REGION Network 3
   RUNG wire#powerrail
      Contact( "FB11_DATA_ALARM_FB_DB".PIW258.QH_ALM )
      wire#w1
      P_Trig( "DB9_P".P2 )
      S_Coil( "Tag_32" )
   END_RUNG
   RUNG wire#powerrail
      Contact( "FB11_DATA_ALARM_FB_DB".PIW258.QL_ALM )
   END_RUNG wire#w1
   // the same network as SCL:
   #_w1 := "FB11_DATA_ALARM_FB_DB".PIW258.QH_ALM OR "FB11_DATA_ALARM_FB_DB".PIW258.QL_ALM;
   #_w2 := #_w1 AND NOT "DB9_P".P2;   // rising edge
   "DB9_P".P2 := #_w1;
   IF #_w2 THEN "Tag_32" := TRUE; END_IF;
END_REGION

REGION Network 4
   RUNG wire#powerrail
      Contact( "FB11_DATA_ALARM_FB_DB".PIW260.QH_ALM )
      wire#w1
      P_Trig( "DB9_P".P3 )
      S_Coil( "Tag_32" )
   END_RUNG
   RUNG wire#powerrail
      Contact( "FB11_DATA_ALARM_FB_DB".PIW260.QL_ALM )
   END_RUNG wire#w1
   // the same network as SCL:
   #_w1 := "FB11_DATA_ALARM_FB_DB".PIW260.QH_ALM OR "FB11_DATA_ALARM_FB_DB".PIW260.QL_ALM;
   #_w2 := #_w1 AND NOT "DB9_P".P3;   // rising edge
   "DB9_P".P3 := #_w1;
   IF #_w2 THEN "Tag_32" := TRUE; END_IF;
END_REGION

REGION Network 5
   RUNG wire#powerrail
      Contact( "FB11_DATA_ALARM_FB_DB".PIW262.QH_ALM )
      wire#w1
      P_Trig( "DB9_P".P4 )
      S_Coil( "Tag_32" )
   END_RUNG
   RUNG wire#powerrail
      Contact( "FB11_DATA_ALARM_FB_DB".PIW262.QL_ALM )
   END_RUNG wire#w1
   // the same network as SCL:
   #_w1 := "FB11_DATA_ALARM_FB_DB".PIW262.QH_ALM OR "FB11_DATA_ALARM_FB_DB".PIW262.QL_ALM;
   #_w2 := #_w1 AND NOT "DB9_P".P4;   // rising edge
   "DB9_P".P4 := #_w1;
   IF #_w2 THEN "Tag_32" := TRUE; END_IF;
END_REGION

REGION Network 6
   RUNG wire#powerrail
      Contact( "FB11_DATA_ALARM_FB_DB".PIW264.QH_ALM )
      wire#w1
      P_Trig( "DB9_P".P5 )
      S_Coil( "Tag_32" )
   END_RUNG
   RUNG wire#powerrail
      Contact( "FB11_DATA_ALARM_FB_DB".PIW264.QL_ALM )
   END_RUNG wire#w1
   // the same network as SCL:
   #_w1 := "FB11_DATA_ALARM_FB_DB".PIW264.QH_ALM OR "FB11_DATA_ALARM_FB_DB".PIW264.QL_ALM;
   #_w2 := #_w1 AND NOT "DB9_P".P5;   // rising edge
   "DB9_P".P5 := #_w1;
   IF #_w2 THEN "Tag_32" := TRUE; END_IF;
END_REGION

REGION Network 7
   RUNG wire#powerrail
      Contact( "FB11_DATA_ALARM_FB_DB".PIW266.QH_ALM )
      wire#w1
      P_Trig( "DB9_P".P6 )
      S_Coil( "Tag_32" )
   END_RUNG
   RUNG wire#powerrail
      Contact( "FB11_DATA_ALARM_FB_DB".PIW266.QL_ALM )
   END_RUNG wire#w1
   // the same network as SCL:
   #_w1 := "FB11_DATA_ALARM_FB_DB".PIW266.QH_ALM OR "FB11_DATA_ALARM_FB_DB".PIW266.QL_ALM;
   #_w2 := #_w1 AND NOT "DB9_P".P6;   // rising edge
   "DB9_P".P6 := #_w1;
   IF #_w2 THEN "Tag_32" := TRUE; END_IF;
END_REGION

REGION Network 8
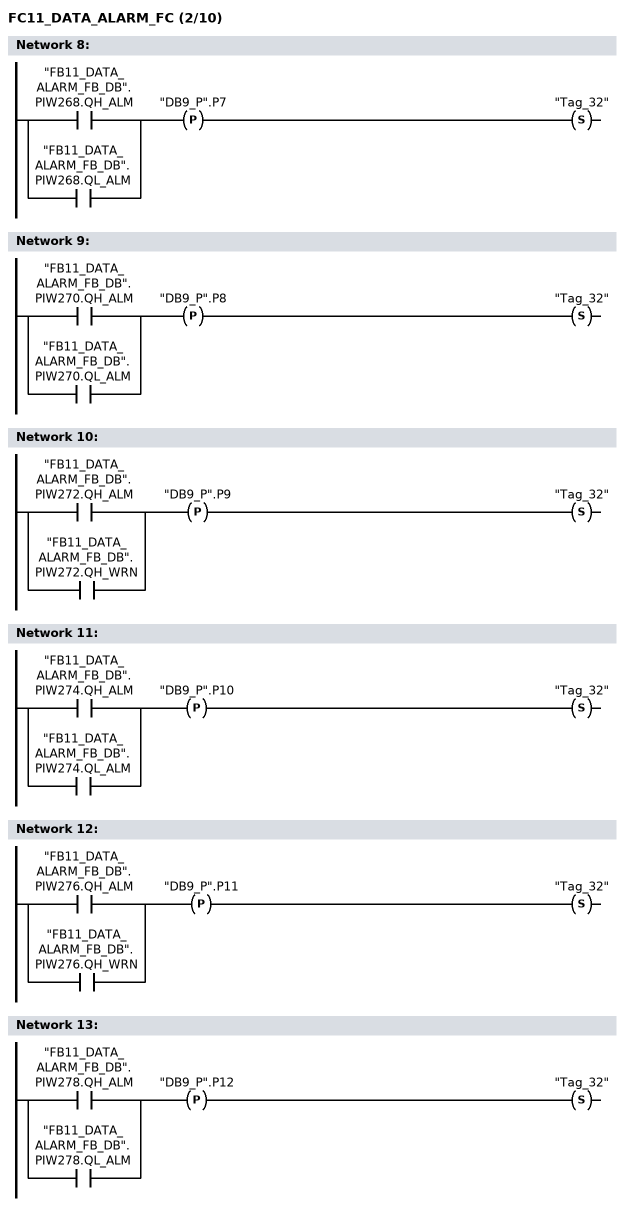
   RUNG wire#powerrail
      Contact( "FB11_DATA_ALARM_FB_DB".PIW268.QH_ALM )
      wire#w1
      P_Trig( "DB9_P".P7 )
      S_Coil( "Tag_32" )
   END_RUNG
   RUNG wire#powerrail
      Contact( "FB11_DATA_ALARM_FB_DB".PIW268.QL_ALM )
   END_RUNG wire#w1
   // the same network as SCL:
   #_w1 := "FB11_DATA_ALARM_FB_DB".PIW268.QH_ALM OR "FB11_DATA_ALARM_FB_DB".PIW268.QL_ALM;
   #_w2 := #_w1 AND NOT "DB9_P".P7;   // rising edge
   "DB9_P".P7 := #_w1;
   IF #_w2 THEN "Tag_32" := TRUE; END_IF;
END_REGION

REGION Network 9
   RUNG wire#powerrail
      Contact( "FB11_DATA_ALARM_FB_DB".PIW270.QH_ALM )
      wire#w1
      P_Trig( "DB9_P".P8 )
      S_Coil( "Tag_32" )
   END_RUNG
   RUNG wire#powerrail
      Contact( "FB11_DATA_ALARM_FB_DB".PIW270.QL_ALM )
   END_RUNG wire#w1
   // the same network as SCL:
   #_w1 := "FB11_DATA_ALARM_FB_DB".PIW270.QH_ALM OR "FB11_DATA_ALARM_FB_DB".PIW270.QL_ALM;
   #_w2 := #_w1 AND NOT "DB9_P".P8;   // rising edge
   "DB9_P".P8 := #_w1;
   IF #_w2 THEN "Tag_32" := TRUE; END_IF;
END_REGION

REGION Network 10
   RUNG wire#powerrail
      Contact( "FB11_DATA_ALARM_FB_DB".PIW272.QH_ALM )
      wire#w1
      P_Trig( "DB9_P".P9 )
      S_Coil( "Tag_32" )
   END_RUNG
   RUNG wire#powerrail
      Contact( "FB11_DATA_ALARM_FB_DB".PIW272.QH_WRN )
   END_RUNG wire#w1
   // the same network as SCL:
   #_w1 := "FB11_DATA_ALARM_FB_DB".PIW272.QH_ALM OR "FB11_DATA_ALARM_FB_DB".PIW272.QH_WRN;
   #_w2 := #_w1 AND NOT "DB9_P".P9;   // rising edge
   "DB9_P".P9 := #_w1;
   IF #_w2 THEN "Tag_32" := TRUE; END_IF;
END_REGION

REGION Network 11
   RUNG wire#powerrail
      Contact( "FB11_DATA_ALARM_FB_DB".PIW274.QH_ALM )
      wire#w1
      P_Trig( "DB9_P".P10 )
      S_Coil( "Tag_32" )
   END_RUNG
   RUNG wire#powerrail
      Contact( "FB11_DATA_ALARM_FB_DB".PIW274.QL_ALM )
   END_RUNG wire#w1
   // the same network as SCL:
   #_w1 := "FB11_DATA_ALARM_FB_DB".PIW274.QH_ALM OR "FB11_DATA_ALARM_FB_DB".PIW274.QL_ALM;
   #_w2 := #_w1 AND NOT "DB9_P".P10;   // rising edge
   "DB9_P".P10 := #_w1;
   IF #_w2 THEN "Tag_32" := TRUE; END_IF;
END_REGION

REGION Network 12
   RUNG wire#powerrail
      Contact( "FB11_DATA_ALARM_FB_DB".PIW276.QH_ALM )
      wire#w1
      P_Trig( "DB9_P".P11 )
      S_Coil( "Tag_32" )
   END_RUNG
   RUNG wire#powerrail
      Contact( "FB11_DATA_ALARM_FB_DB".PIW276.QH_WRN )
   END_RUNG wire#w1
   // the same network as SCL:
   #_w1 := "FB11_DATA_ALARM_FB_DB".PIW276.QH_ALM OR "FB11_DATA_ALARM_FB_DB".PIW276.QH_WRN;
   #_w2 := #_w1 AND NOT "DB9_P".P11;   // rising edge
   "DB9_P".P11 := #_w1;
   IF #_w2 THEN "Tag_32" := TRUE; END_IF;
END_REGION

REGION Network 13
   RUNG wire#powerrail
      Contact( "FB11_DATA_ALARM_FB_DB".PIW278.QH_ALM )
      wire#w1
      P_Trig( "DB9_P".P12 )
      S_Coil( "Tag_32" )
   END_RUNG
   RUNG wire#powerrail
      Contact( "FB11_DATA_ALARM_FB_DB".PIW278.QL_ALM )
   END_RUNG wire#w1
   // the same network as SCL:
   #_w1 := "FB11_DATA_ALARM_FB_DB".PIW278.QH_ALM OR "FB11_DATA_ALARM_FB_DB".PIW278.QL_ALM;
   #_w2 := #_w1 AND NOT "DB9_P".P12;   // rising edge
   "DB9_P".P12 := #_w1;
   IF #_w2 THEN "Tag_32" := TRUE; END_IF;
END_REGION

REGION Network 14
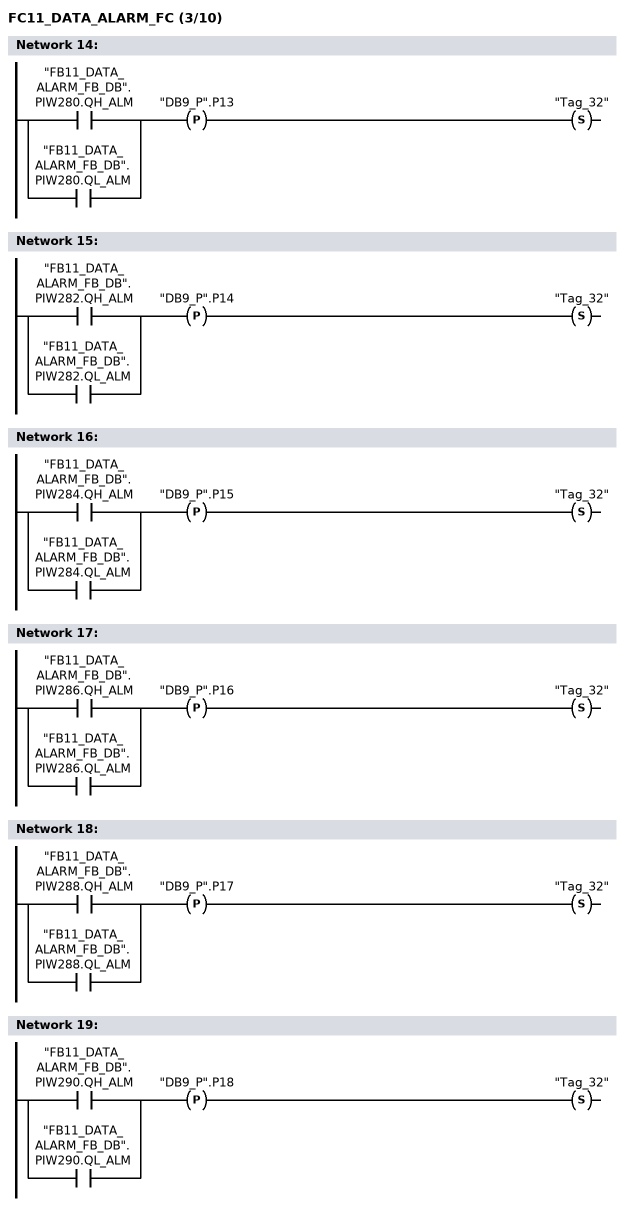
   RUNG wire#powerrail
      Contact( "FB11_DATA_ALARM_FB_DB".PIW280.QH_ALM )
      wire#w1
      P_Trig( "DB9_P".P13 )
      S_Coil( "Tag_32" )
   END_RUNG
   RUNG wire#powerrail
      Contact( "FB11_DATA_ALARM_FB_DB".PIW280.QL_ALM )
   END_RUNG wire#w1
   // the same network as SCL:
   #_w1 := "FB11_DATA_ALARM_FB_DB".PIW280.QH_ALM OR "FB11_DATA_ALARM_FB_DB".PIW280.QL_ALM;
   #_w2 := #_w1 AND NOT "DB9_P".P13;   // rising edge
   "DB9_P".P13 := #_w1;
   IF #_w2 THEN "Tag_32" := TRUE; END_IF;
END_REGION

REGION Network 15
   RUNG wire#powerrail
      Contact( "FB11_DATA_ALARM_FB_DB".PIW282.QH_ALM )
      wire#w1
      P_Trig( "DB9_P".P14 )
      S_Coil( "Tag_32" )
   END_RUNG
   RUNG wire#powerrail
      Contact( "FB11_DATA_ALARM_FB_DB".PIW282.QL_ALM )
   END_RUNG wire#w1
   // the same network as SCL:
   #_w1 := "FB11_DATA_ALARM_FB_DB".PIW282.QH_ALM OR "FB11_DATA_ALARM_FB_DB".PIW282.QL_ALM;
   #_w2 := #_w1 AND NOT "DB9_P".P14;   // rising edge
   "DB9_P".P14 := #_w1;
   IF #_w2 THEN "Tag_32" := TRUE; END_IF;
END_REGION

REGION Network 16
   RUNG wire#powerrail
      Contact( "FB11_DATA_ALARM_FB_DB".PIW284.QH_ALM )
      wire#w1
      P_Trig( "DB9_P".P15 )
      S_Coil( "Tag_32" )
   END_RUNG
   RUNG wire#powerrail
      Contact( "FB11_DATA_ALARM_FB_DB".PIW284.QL_ALM )
   END_RUNG wire#w1
   // the same network as SCL:
   #_w1 := "FB11_DATA_ALARM_FB_DB".PIW284.QH_ALM OR "FB11_DATA_ALARM_FB_DB".PIW284.QL_ALM;
   #_w2 := #_w1 AND NOT "DB9_P".P15;   // rising edge
   "DB9_P".P15 := #_w1;
   IF #_w2 THEN "Tag_32" := TRUE; END_IF;
END_REGION

REGION Network 17
   RUNG wire#powerrail
      Contact( "FB11_DATA_ALARM_FB_DB".PIW286.QH_ALM )
      wire#w1
      P_Trig( "DB9_P".P16 )
      S_Coil( "Tag_32" )
   END_RUNG
   RUNG wire#powerrail
      Contact( "FB11_DATA_ALARM_FB_DB".PIW286.QL_ALM )
   END_RUNG wire#w1
   // the same network as SCL:
   #_w1 := "FB11_DATA_ALARM_FB_DB".PIW286.QH_ALM OR "FB11_DATA_ALARM_FB_DB".PIW286.QL_ALM;
   #_w2 := #_w1 AND NOT "DB9_P".P16;   // rising edge
   "DB9_P".P16 := #_w1;
   IF #_w2 THEN "Tag_32" := TRUE; END_IF;
END_REGION

REGION Network 18
   RUNG wire#powerrail
      Contact( "FB11_DATA_ALARM_FB_DB".PIW288.QH_ALM )
      wire#w1
      P_Trig( "DB9_P".P17 )
      S_Coil( "Tag_32" )
   END_RUNG
   RUNG wire#powerrail
      Contact( "FB11_DATA_ALARM_FB_DB".PIW288.QL_ALM )
   END_RUNG wire#w1
   // the same network as SCL:
   #_w1 := "FB11_DATA_ALARM_FB_DB".PIW288.QH_ALM OR "FB11_DATA_ALARM_FB_DB".PIW288.QL_ALM;
   #_w2 := #_w1 AND NOT "DB9_P".P17;   // rising edge
   "DB9_P".P17 := #_w1;
   IF #_w2 THEN "Tag_32" := TRUE; END_IF;
END_REGION

REGION Network 19
   RUNG wire#powerrail
      Contact( "FB11_DATA_ALARM_FB_DB".PIW290.QH_ALM )
      wire#w1
      P_Trig( "DB9_P".P18 )
      S_Coil( "Tag_32" )
   END_RUNG
   RUNG wire#powerrail
      Contact( "FB11_DATA_ALARM_FB_DB".PIW290.QL_ALM )
   END_RUNG wire#w1
   // the same network as SCL:
   #_w1 := "FB11_DATA_ALARM_FB_DB".PIW290.QH_ALM OR "FB11_DATA_ALARM_FB_DB".PIW290.QL_ALM;
   #_w2 := #_w1 AND NOT "DB9_P".P18;   // rising edge
   "DB9_P".P18 := #_w1;
   IF #_w2 THEN "Tag_32" := TRUE; END_IF;
END_REGION

REGION Network 20
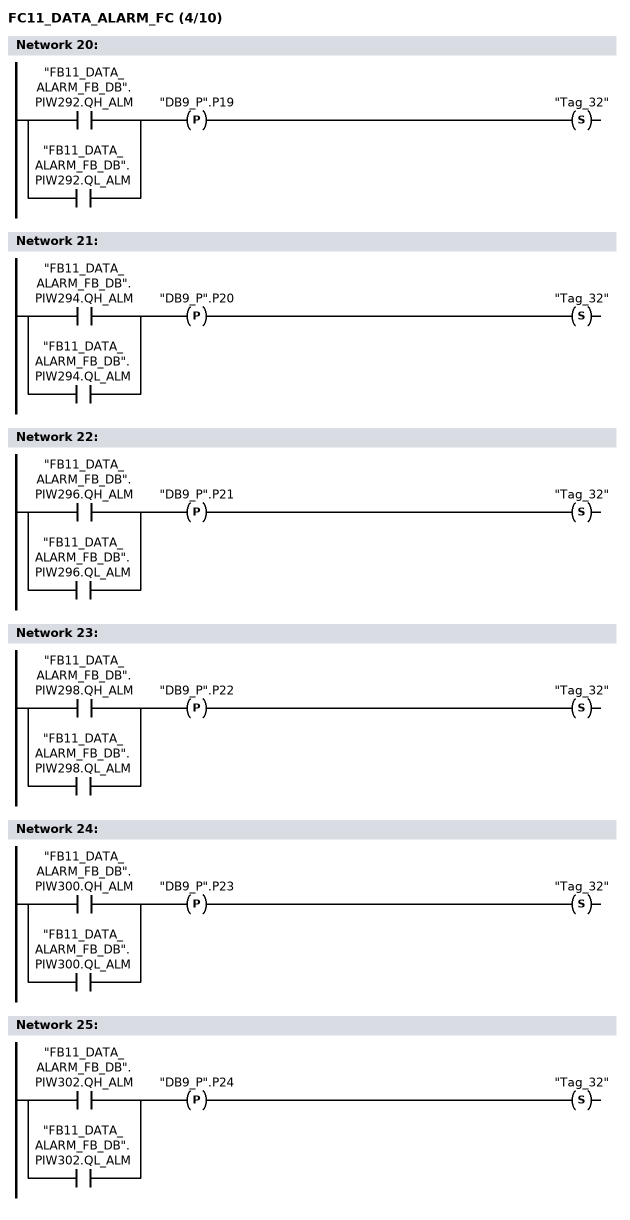
   RUNG wire#powerrail
      Contact( "FB11_DATA_ALARM_FB_DB".PIW292.QH_ALM )
      wire#w1
      P_Trig( "DB9_P".P19 )
      S_Coil( "Tag_32" )
   END_RUNG
   RUNG wire#powerrail
      Contact( "FB11_DATA_ALARM_FB_DB".PIW292.QL_ALM )
   END_RUNG wire#w1
   // the same network as SCL:
   #_w1 := "FB11_DATA_ALARM_FB_DB".PIW292.QH_ALM OR "FB11_DATA_ALARM_FB_DB".PIW292.QL_ALM;
   #_w2 := #_w1 AND NOT "DB9_P".P19;   // rising edge
   "DB9_P".P19 := #_w1;
   IF #_w2 THEN "Tag_32" := TRUE; END_IF;
END_REGION

REGION Network 21
   RUNG wire#powerrail
      Contact( "FB11_DATA_ALARM_FB_DB".PIW294.QH_ALM )
      wire#w1
      P_Trig( "DB9_P".P20 )
      S_Coil( "Tag_32" )
   END_RUNG
   RUNG wire#powerrail
      Contact( "FB11_DATA_ALARM_FB_DB".PIW294.QL_ALM )
   END_RUNG wire#w1
   // the same network as SCL:
   #_w1 := "FB11_DATA_ALARM_FB_DB".PIW294.QH_ALM OR "FB11_DATA_ALARM_FB_DB".PIW294.QL_ALM;
   #_w2 := #_w1 AND NOT "DB9_P".P20;   // rising edge
   "DB9_P".P20 := #_w1;
   IF #_w2 THEN "Tag_32" := TRUE; END_IF;
END_REGION

REGION Network 22
   RUNG wire#powerrail
      Contact( "FB11_DATA_ALARM_FB_DB".PIW296.QH_ALM )
      wire#w1
      P_Trig( "DB9_P".P21 )
      S_Coil( "Tag_32" )
   END_RUNG
   RUNG wire#powerrail
      Contact( "FB11_DATA_ALARM_FB_DB".PIW296.QL_ALM )
   END_RUNG wire#w1
   // the same network as SCL:
   #_w1 := "FB11_DATA_ALARM_FB_DB".PIW296.QH_ALM OR "FB11_DATA_ALARM_FB_DB".PIW296.QL_ALM;
   #_w2 := #_w1 AND NOT "DB9_P".P21;   // rising edge
   "DB9_P".P21 := #_w1;
   IF #_w2 THEN "Tag_32" := TRUE; END_IF;
END_REGION

REGION Network 23
   RUNG wire#powerrail
      Contact( "FB11_DATA_ALARM_FB_DB".PIW298.QH_ALM )
      wire#w1
      P_Trig( "DB9_P".P22 )
      S_Coil( "Tag_32" )
   END_RUNG
   RUNG wire#powerrail
      Contact( "FB11_DATA_ALARM_FB_DB".PIW298.QL_ALM )
   END_RUNG wire#w1
   // the same network as SCL:
   #_w1 := "FB11_DATA_ALARM_FB_DB".PIW298.QH_ALM OR "FB11_DATA_ALARM_FB_DB".PIW298.QL_ALM;
   #_w2 := #_w1 AND NOT "DB9_P".P22;   // rising edge
   "DB9_P".P22 := #_w1;
   IF #_w2 THEN "Tag_32" := TRUE; END_IF;
END_REGION

REGION Network 24
   RUNG wire#powerrail
      Contact( "FB11_DATA_ALARM_FB_DB".PIW300.QH_ALM )
      wire#w1
      P_Trig( "DB9_P".P23 )
      S_Coil( "Tag_32" )
   END_RUNG
   RUNG wire#powerrail
      Contact( "FB11_DATA_ALARM_FB_DB".PIW300.QL_ALM )
   END_RUNG wire#w1
   // the same network as SCL:
   #_w1 := "FB11_DATA_ALARM_FB_DB".PIW300.QH_ALM OR "FB11_DATA_ALARM_FB_DB".PIW300.QL_ALM;
   #_w2 := #_w1 AND NOT "DB9_P".P23;   // rising edge
   "DB9_P".P23 := #_w1;
   IF #_w2 THEN "Tag_32" := TRUE; END_IF;
END_REGION

REGION Network 25
   RUNG wire#powerrail
      Contact( "FB11_DATA_ALARM_FB_DB".PIW302.QH_ALM )
      wire#w1
      P_Trig( "DB9_P".P24 )
      S_Coil( "Tag_32" )
   END_RUNG
   RUNG wire#powerrail
      Contact( "FB11_DATA_ALARM_FB_DB".PIW302.QL_ALM )
   END_RUNG wire#w1
   // the same network as SCL:
   #_w1 := "FB11_DATA_ALARM_FB_DB".PIW302.QH_ALM OR "FB11_DATA_ALARM_FB_DB".PIW302.QL_ALM;
   #_w2 := #_w1 AND NOT "DB9_P".P24;   // rising edge
   "DB9_P".P24 := #_w1;
   IF #_w2 THEN "Tag_32" := TRUE; END_IF;
END_REGION

REGION Network 26
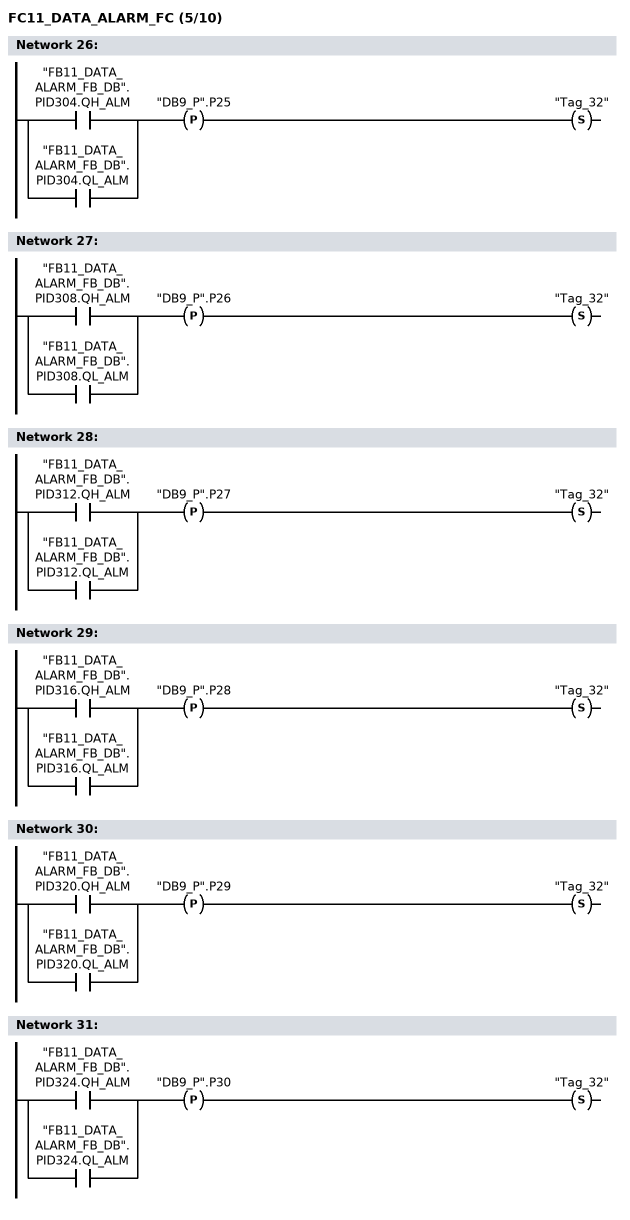
   RUNG wire#powerrail
      Contact( "FB11_DATA_ALARM_FB_DB".PID304.QH_ALM )
      wire#w1
      P_Trig( "DB9_P".P25 )
      S_Coil( "Tag_32" )
   END_RUNG
   RUNG wire#powerrail
      Contact( "FB11_DATA_ALARM_FB_DB".PID304.QL_ALM )
   END_RUNG wire#w1
   // the same network as SCL:
   #_w1 := "FB11_DATA_ALARM_FB_DB".PID304.QH_ALM OR "FB11_DATA_ALARM_FB_DB".PID304.QL_ALM;
   #_w2 := #_w1 AND NOT "DB9_P".P25;   // rising edge
   "DB9_P".P25 := #_w1;
   IF #_w2 THEN "Tag_32" := TRUE; END_IF;
END_REGION

REGION Network 27
   RUNG wire#powerrail
      Contact( "FB11_DATA_ALARM_FB_DB".PID308.QH_ALM )
      wire#w1
      P_Trig( "DB9_P".P26 )
      S_Coil( "Tag_32" )
   END_RUNG
   RUNG wire#powerrail
      Contact( "FB11_DATA_ALARM_FB_DB".PID308.QL_ALM )
   END_RUNG wire#w1
   // the same network as SCL:
   #_w1 := "FB11_DATA_ALARM_FB_DB".PID308.QH_ALM OR "FB11_DATA_ALARM_FB_DB".PID308.QL_ALM;
   #_w2 := #_w1 AND NOT "DB9_P".P26;   // rising edge
   "DB9_P".P26 := #_w1;
   IF #_w2 THEN "Tag_32" := TRUE; END_IF;
END_REGION

REGION Network 28
   RUNG wire#powerrail
      Contact( "FB11_DATA_ALARM_FB_DB".PID312.QH_ALM )
      wire#w1
      P_Trig( "DB9_P".P27 )
      S_Coil( "Tag_32" )
   END_RUNG
   RUNG wire#powerrail
      Contact( "FB11_DATA_ALARM_FB_DB".PID312.QL_ALM )
   END_RUNG wire#w1
   // the same network as SCL:
   #_w1 := "FB11_DATA_ALARM_FB_DB".PID312.QH_ALM OR "FB11_DATA_ALARM_FB_DB".PID312.QL_ALM;
   #_w2 := #_w1 AND NOT "DB9_P".P27;   // rising edge
   "DB9_P".P27 := #_w1;
   IF #_w2 THEN "Tag_32" := TRUE; END_IF;
END_REGION

REGION Network 29
   RUNG wire#powerrail
      Contact( "FB11_DATA_ALARM_FB_DB".PID316.QH_ALM )
      wire#w1
      P_Trig( "DB9_P".P28 )
      S_Coil( "Tag_32" )
   END_RUNG
   RUNG wire#powerrail
      Contact( "FB11_DATA_ALARM_FB_DB".PID316.QL_ALM )
   END_RUNG wire#w1
   // the same network as SCL:
   #_w1 := "FB11_DATA_ALARM_FB_DB".PID316.QH_ALM OR "FB11_DATA_ALARM_FB_DB".PID316.QL_ALM;
   #_w2 := #_w1 AND NOT "DB9_P".P28;   // rising edge
   "DB9_P".P28 := #_w1;
   IF #_w2 THEN "Tag_32" := TRUE; END_IF;
END_REGION

REGION Network 30
   RUNG wire#powerrail
      Contact( "FB11_DATA_ALARM_FB_DB".PID320.QH_ALM )
      wire#w1
      P_Trig( "DB9_P".P29 )
      S_Coil( "Tag_32" )
   END_RUNG
   RUNG wire#powerrail
      Contact( "FB11_DATA_ALARM_FB_DB".PID320.QL_ALM )
   END_RUNG wire#w1
   // the same network as SCL:
   #_w1 := "FB11_DATA_ALARM_FB_DB".PID320.QH_ALM OR "FB11_DATA_ALARM_FB_DB".PID320.QL_ALM;
   #_w2 := #_w1 AND NOT "DB9_P".P29;   // rising edge
   "DB9_P".P29 := #_w1;
   IF #_w2 THEN "Tag_32" := TRUE; END_IF;
END_REGION

REGION Network 31
   RUNG wire#powerrail
      Contact( "FB11_DATA_ALARM_FB_DB".PID324.QH_ALM )
      wire#w1
      P_Trig( "DB9_P".P30 )
      S_Coil( "Tag_32" )
   END_RUNG
   RUNG wire#powerrail
      Contact( "FB11_DATA_ALARM_FB_DB".PID324.QL_ALM )
   END_RUNG wire#w1
   // the same network as SCL:
   #_w1 := "FB11_DATA_ALARM_FB_DB".PID324.QH_ALM OR "FB11_DATA_ALARM_FB_DB".PID324.QL_ALM;
   #_w2 := #_w1 AND NOT "DB9_P".P30;   // rising edge
   "DB9_P".P30 := #_w1;
   IF #_w2 THEN "Tag_32" := TRUE; END_IF;
END_REGION

REGION Network 32
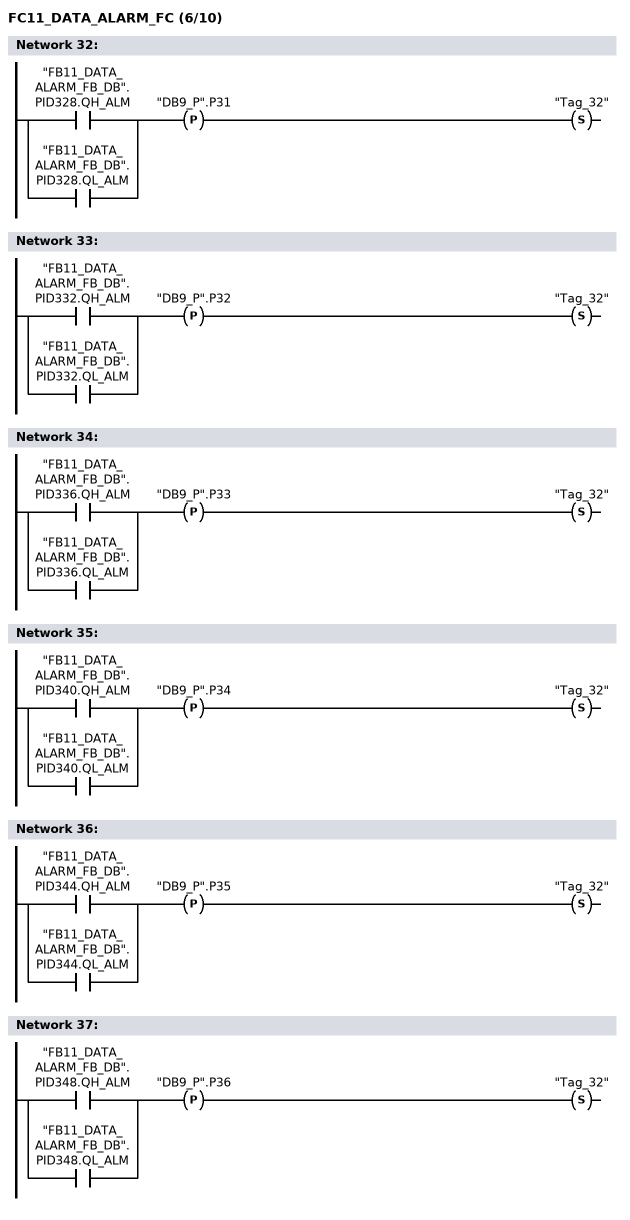
   RUNG wire#powerrail
      Contact( "FB11_DATA_ALARM_FB_DB".PID328.QH_ALM )
      wire#w1
      P_Trig( "DB9_P".P31 )
      S_Coil( "Tag_32" )
   END_RUNG
   RUNG wire#powerrail
      Contact( "FB11_DATA_ALARM_FB_DB".PID328.QL_ALM )
   END_RUNG wire#w1
   // the same network as SCL:
   #_w1 := "FB11_DATA_ALARM_FB_DB".PID328.QH_ALM OR "FB11_DATA_ALARM_FB_DB".PID328.QL_ALM;
   #_w2 := #_w1 AND NOT "DB9_P".P31;   // rising edge
   "DB9_P".P31 := #_w1;
   IF #_w2 THEN "Tag_32" := TRUE; END_IF;
END_REGION

REGION Network 33
   RUNG wire#powerrail
      Contact( "FB11_DATA_ALARM_FB_DB".PID332.QH_ALM )
      wire#w1
      P_Trig( "DB9_P".P32 )
      S_Coil( "Tag_32" )
   END_RUNG
   RUNG wire#powerrail
      Contact( "FB11_DATA_ALARM_FB_DB".PID332.QL_ALM )
   END_RUNG wire#w1
   // the same network as SCL:
   #_w1 := "FB11_DATA_ALARM_FB_DB".PID332.QH_ALM OR "FB11_DATA_ALARM_FB_DB".PID332.QL_ALM;
   #_w2 := #_w1 AND NOT "DB9_P".P32;   // rising edge
   "DB9_P".P32 := #_w1;
   IF #_w2 THEN "Tag_32" := TRUE; END_IF;
END_REGION

REGION Network 34
   RUNG wire#powerrail
      Contact( "FB11_DATA_ALARM_FB_DB".PID336.QH_ALM )
      wire#w1
      P_Trig( "DB9_P".P33 )
      S_Coil( "Tag_32" )
   END_RUNG
   RUNG wire#powerrail
      Contact( "FB11_DATA_ALARM_FB_DB".PID336.QL_ALM )
   END_RUNG wire#w1
   // the same network as SCL:
   #_w1 := "FB11_DATA_ALARM_FB_DB".PID336.QH_ALM OR "FB11_DATA_ALARM_FB_DB".PID336.QL_ALM;
   #_w2 := #_w1 AND NOT "DB9_P".P33;   // rising edge
   "DB9_P".P33 := #_w1;
   IF #_w2 THEN "Tag_32" := TRUE; END_IF;
END_REGION

REGION Network 35
   RUNG wire#powerrail
      Contact( "FB11_DATA_ALARM_FB_DB".PID340.QH_ALM )
      wire#w1
      P_Trig( "DB9_P".P34 )
      S_Coil( "Tag_32" )
   END_RUNG
   RUNG wire#powerrail
      Contact( "FB11_DATA_ALARM_FB_DB".PID340.QL_ALM )
   END_RUNG wire#w1
   // the same network as SCL:
   #_w1 := "FB11_DATA_ALARM_FB_DB".PID340.QH_ALM OR "FB11_DATA_ALARM_FB_DB".PID340.QL_ALM;
   #_w2 := #_w1 AND NOT "DB9_P".P34;   // rising edge
   "DB9_P".P34 := #_w1;
   IF #_w2 THEN "Tag_32" := TRUE; END_IF;
END_REGION

REGION Network 36
   RUNG wire#powerrail
      Contact( "FB11_DATA_ALARM_FB_DB".PID344.QH_ALM )
      wire#w1
      P_Trig( "DB9_P".P35 )
      S_Coil( "Tag_32" )
   END_RUNG
   RUNG wire#powerrail
      Contact( "FB11_DATA_ALARM_FB_DB".PID344.QL_ALM )
   END_RUNG wire#w1
   // the same network as SCL:
   #_w1 := "FB11_DATA_ALARM_FB_DB".PID344.QH_ALM OR "FB11_DATA_ALARM_FB_DB".PID344.QL_ALM;
   #_w2 := #_w1 AND NOT "DB9_P".P35;   // rising edge
   "DB9_P".P35 := #_w1;
   IF #_w2 THEN "Tag_32" := TRUE; END_IF;
END_REGION

REGION Network 37
   RUNG wire#powerrail
      Contact( "FB11_DATA_ALARM_FB_DB".PID348.QH_ALM )
      wire#w1
      P_Trig( "DB9_P".P36 )
      S_Coil( "Tag_32" )
   END_RUNG
   RUNG wire#powerrail
      Contact( "FB11_DATA_ALARM_FB_DB".PID348.QL_ALM )
   END_RUNG wire#w1
   // the same network as SCL:
   #_w1 := "FB11_DATA_ALARM_FB_DB".PID348.QH_ALM OR "FB11_DATA_ALARM_FB_DB".PID348.QL_ALM;
   #_w2 := #_w1 AND NOT "DB9_P".P36;   // rising edge
   "DB9_P".P36 := #_w1;
   IF #_w2 THEN "Tag_32" := TRUE; END_IF;
END_REGION

REGION Network 38
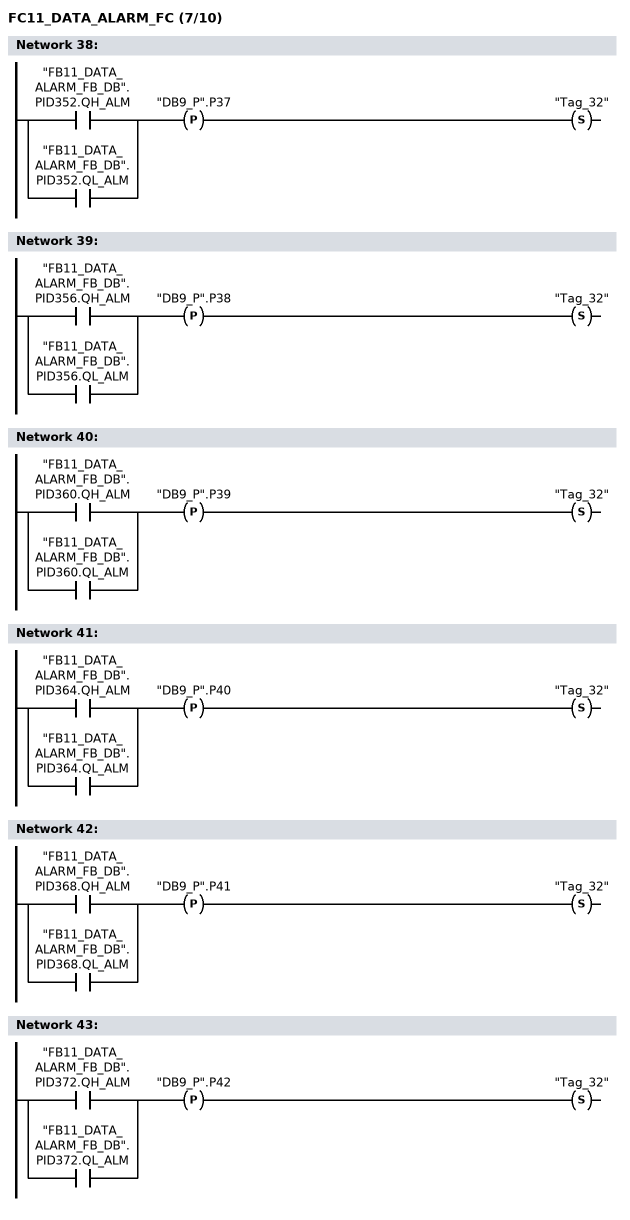
   RUNG wire#powerrail
      Contact( "FB11_DATA_ALARM_FB_DB".PID352.QH_ALM )
      wire#w1
      P_Trig( "DB9_P".P37 )
      S_Coil( "Tag_32" )
   END_RUNG
   RUNG wire#powerrail
      Contact( "FB11_DATA_ALARM_FB_DB".PID352.QL_ALM )
   END_RUNG wire#w1
   // the same network as SCL:
   #_w1 := "FB11_DATA_ALARM_FB_DB".PID352.QH_ALM OR "FB11_DATA_ALARM_FB_DB".PID352.QL_ALM;
   #_w2 := #_w1 AND NOT "DB9_P".P37;   // rising edge
   "DB9_P".P37 := #_w1;
   IF #_w2 THEN "Tag_32" := TRUE; END_IF;
END_REGION

REGION Network 39
   RUNG wire#powerrail
      Contact( "FB11_DATA_ALARM_FB_DB".PID356.QH_ALM )
      wire#w1
      P_Trig( "DB9_P".P38 )
      S_Coil( "Tag_32" )
   END_RUNG
   RUNG wire#powerrail
      Contact( "FB11_DATA_ALARM_FB_DB".PID356.QL_ALM )
   END_RUNG wire#w1
   // the same network as SCL:
   #_w1 := "FB11_DATA_ALARM_FB_DB".PID356.QH_ALM OR "FB11_DATA_ALARM_FB_DB".PID356.QL_ALM;
   #_w2 := #_w1 AND NOT "DB9_P".P38;   // rising edge
   "DB9_P".P38 := #_w1;
   IF #_w2 THEN "Tag_32" := TRUE; END_IF;
END_REGION

REGION Network 40
   RUNG wire#powerrail
      Contact( "FB11_DATA_ALARM_FB_DB".PID360.QH_ALM )
      wire#w1
      P_Trig( "DB9_P".P39 )
      S_Coil( "Tag_32" )
   END_RUNG
   RUNG wire#powerrail
      Contact( "FB11_DATA_ALARM_FB_DB".PID360.QL_ALM )
   END_RUNG wire#w1
   // the same network as SCL:
   #_w1 := "FB11_DATA_ALARM_FB_DB".PID360.QH_ALM OR "FB11_DATA_ALARM_FB_DB".PID360.QL_ALM;
   #_w2 := #_w1 AND NOT "DB9_P".P39;   // rising edge
   "DB9_P".P39 := #_w1;
   IF #_w2 THEN "Tag_32" := TRUE; END_IF;
END_REGION

REGION Network 41
   RUNG wire#powerrail
      Contact( "FB11_DATA_ALARM_FB_DB".PID364.QH_ALM )
      wire#w1
      P_Trig( "DB9_P".P40 )
      S_Coil( "Tag_32" )
   END_RUNG
   RUNG wire#powerrail
      Contact( "FB11_DATA_ALARM_FB_DB".PID364.QL_ALM )
   END_RUNG wire#w1
   // the same network as SCL:
   #_w1 := "FB11_DATA_ALARM_FB_DB".PID364.QH_ALM OR "FB11_DATA_ALARM_FB_DB".PID364.QL_ALM;
   #_w2 := #_w1 AND NOT "DB9_P".P40;   // rising edge
   "DB9_P".P40 := #_w1;
   IF #_w2 THEN "Tag_32" := TRUE; END_IF;
END_REGION

REGION Network 42
   RUNG wire#powerrail
      Contact( "FB11_DATA_ALARM_FB_DB".PID368.QH_ALM )
      wire#w1
      P_Trig( "DB9_P".P41 )
      S_Coil( "Tag_32" )
   END_RUNG
   RUNG wire#powerrail
      Contact( "FB11_DATA_ALARM_FB_DB".PID368.QL_ALM )
   END_RUNG wire#w1
   // the same network as SCL:
   #_w1 := "FB11_DATA_ALARM_FB_DB".PID368.QH_ALM OR "FB11_DATA_ALARM_FB_DB".PID368.QL_ALM;
   #_w2 := #_w1 AND NOT "DB9_P".P41;   // rising edge
   "DB9_P".P41 := #_w1;
   IF #_w2 THEN "Tag_32" := TRUE; END_IF;
END_REGION

REGION Network 43
   RUNG wire#powerrail
      Contact( "FB11_DATA_ALARM_FB_DB".PID372.QH_ALM )
      wire#w1
      P_Trig( "DB9_P".P42 )
      S_Coil( "Tag_32" )
   END_RUNG
   RUNG wire#powerrail
      Contact( "FB11_DATA_ALARM_FB_DB".PID372.QL_ALM )
   END_RUNG wire#w1
   // the same network as SCL:
   #_w1 := "FB11_DATA_ALARM_FB_DB".PID372.QH_ALM OR "FB11_DATA_ALARM_FB_DB".PID372.QL_ALM;
   #_w2 := #_w1 AND NOT "DB9_P".P42;   // rising edge
   "DB9_P".P42 := #_w1;
   IF #_w2 THEN "Tag_32" := TRUE; END_IF;
END_REGION

REGION Network 44
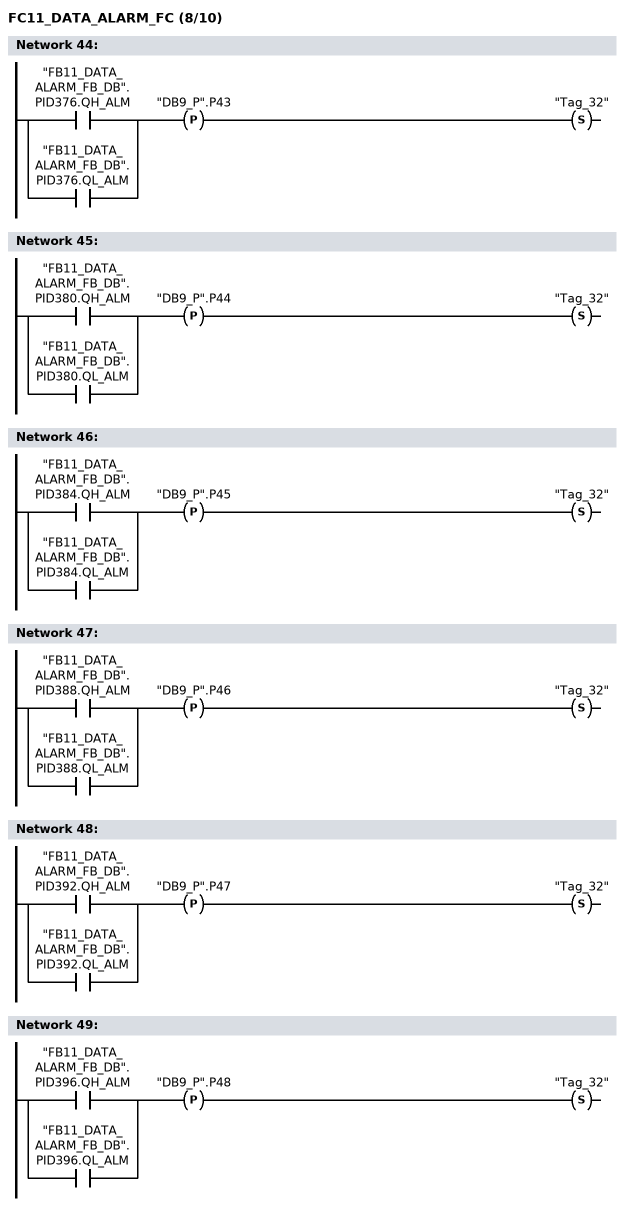
   RUNG wire#powerrail
      Contact( "FB11_DATA_ALARM_FB_DB".PID376.QH_ALM )
      wire#w1
      P_Trig( "DB9_P".P43 )
      S_Coil( "Tag_32" )
   END_RUNG
   RUNG wire#powerrail
      Contact( "FB11_DATA_ALARM_FB_DB".PID376.QL_ALM )
   END_RUNG wire#w1
   // the same network as SCL:
   #_w1 := "FB11_DATA_ALARM_FB_DB".PID376.QH_ALM OR "FB11_DATA_ALARM_FB_DB".PID376.QL_ALM;
   #_w2 := #_w1 AND NOT "DB9_P".P43;   // rising edge
   "DB9_P".P43 := #_w1;
   IF #_w2 THEN "Tag_32" := TRUE; END_IF;
END_REGION

REGION Network 45
   RUNG wire#powerrail
      Contact( "FB11_DATA_ALARM_FB_DB".PID380.QH_ALM )
      wire#w1
      P_Trig( "DB9_P".P44 )
      S_Coil( "Tag_32" )
   END_RUNG
   RUNG wire#powerrail
      Contact( "FB11_DATA_ALARM_FB_DB".PID380.QL_ALM )
   END_RUNG wire#w1
   // the same network as SCL:
   #_w1 := "FB11_DATA_ALARM_FB_DB".PID380.QH_ALM OR "FB11_DATA_ALARM_FB_DB".PID380.QL_ALM;
   #_w2 := #_w1 AND NOT "DB9_P".P44;   // rising edge
   "DB9_P".P44 := #_w1;
   IF #_w2 THEN "Tag_32" := TRUE; END_IF;
END_REGION

REGION Network 46
   RUNG wire#powerrail
      Contact( "FB11_DATA_ALARM_FB_DB".PID384.QH_ALM )
      wire#w1
      P_Trig( "DB9_P".P45 )
      S_Coil( "Tag_32" )
   END_RUNG
   RUNG wire#powerrail
      Contact( "FB11_DATA_ALARM_FB_DB".PID384.QL_ALM )
   END_RUNG wire#w1
   // the same network as SCL:
   #_w1 := "FB11_DATA_ALARM_FB_DB".PID384.QH_ALM OR "FB11_DATA_ALARM_FB_DB".PID384.QL_ALM;
   #_w2 := #_w1 AND NOT "DB9_P".P45;   // rising edge
   "DB9_P".P45 := #_w1;
   IF #_w2 THEN "Tag_32" := TRUE; END_IF;
END_REGION

REGION Network 47
   RUNG wire#powerrail
      Contact( "FB11_DATA_ALARM_FB_DB".PID388.QH_ALM )
      wire#w1
      P_Trig( "DB9_P".P46 )
      S_Coil( "Tag_32" )
   END_RUNG
   RUNG wire#powerrail
      Contact( "FB11_DATA_ALARM_FB_DB".PID388.QL_ALM )
   END_RUNG wire#w1
   // the same network as SCL:
   #_w1 := "FB11_DATA_ALARM_FB_DB".PID388.QH_ALM OR "FB11_DATA_ALARM_FB_DB".PID388.QL_ALM;
   #_w2 := #_w1 AND NOT "DB9_P".P46;   // rising edge
   "DB9_P".P46 := #_w1;
   IF #_w2 THEN "Tag_32" := TRUE; END_IF;
END_REGION

REGION Network 48
   RUNG wire#powerrail
      Contact( "FB11_DATA_ALARM_FB_DB".PID392.QH_ALM )
      wire#w1
      P_Trig( "DB9_P".P47 )
      S_Coil( "Tag_32" )
   END_RUNG
   RUNG wire#powerrail
      Contact( "FB11_DATA_ALARM_FB_DB".PID392.QL_ALM )
   END_RUNG wire#w1
   // the same network as SCL:
   #_w1 := "FB11_DATA_ALARM_FB_DB".PID392.QH_ALM OR "FB11_DATA_ALARM_FB_DB".PID392.QL_ALM;
   #_w2 := #_w1 AND NOT "DB9_P".P47;   // rising edge
   "DB9_P".P47 := #_w1;
   IF #_w2 THEN "Tag_32" := TRUE; END_IF;
END_REGION

REGION Network 49
   RUNG wire#powerrail
      Contact( "FB11_DATA_ALARM_FB_DB".PID396.QH_ALM )
      wire#w1
      P_Trig( "DB9_P".P48 )
      S_Coil( "Tag_32" )
   END_RUNG
   RUNG wire#powerrail
      Contact( "FB11_DATA_ALARM_FB_DB".PID396.QL_ALM )
   END_RUNG wire#w1
   // the same network as SCL:
   #_w1 := "FB11_DATA_ALARM_FB_DB".PID396.QH_ALM OR "FB11_DATA_ALARM_FB_DB".PID396.QL_ALM;
   #_w2 := #_w1 AND NOT "DB9_P".P48;   // rising edge
   "DB9_P".P48 := #_w1;
   IF #_w2 THEN "Tag_32" := TRUE; END_IF;
END_REGION

REGION Network 50
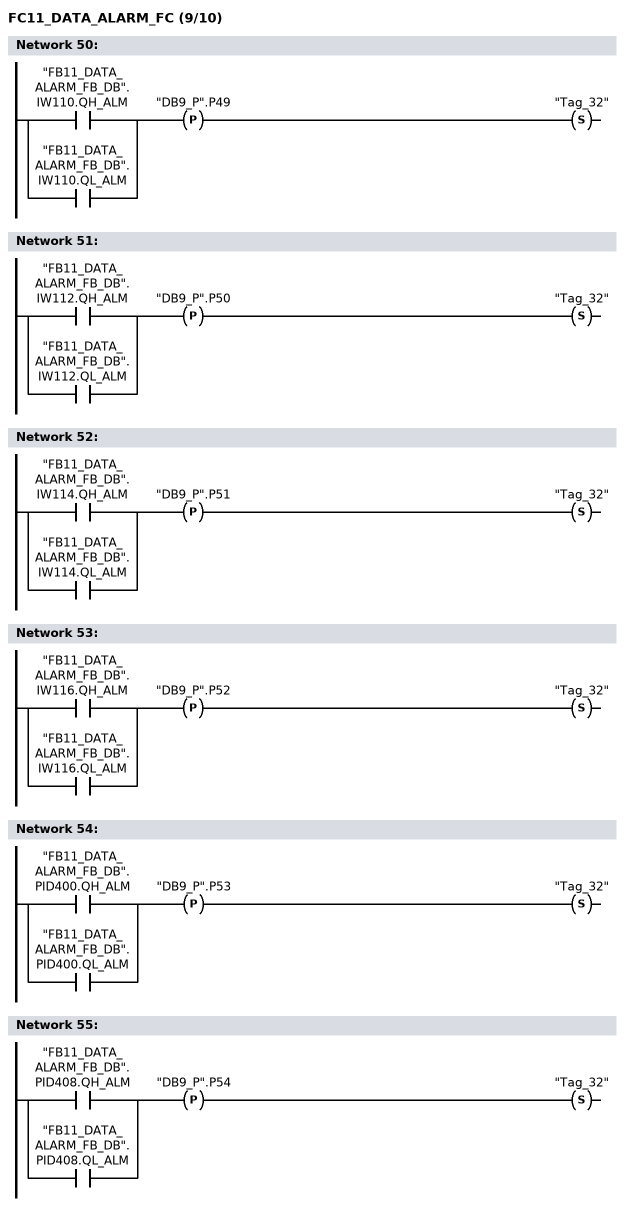
   RUNG wire#powerrail
      Contact( "FB11_DATA_ALARM_FB_DB".IW110.QH_ALM )
      wire#w1
      P_Trig( "DB9_P".P49 )
      S_Coil( "Tag_32" )
   END_RUNG
   RUNG wire#powerrail
      Contact( "FB11_DATA_ALARM_FB_DB".IW110.QL_ALM )
   END_RUNG wire#w1
   // the same network as SCL:
   #_w1 := "FB11_DATA_ALARM_FB_DB".IW110.QH_ALM OR "FB11_DATA_ALARM_FB_DB".IW110.QL_ALM;
   #_w2 := #_w1 AND NOT "DB9_P".P49;   // rising edge
   "DB9_P".P49 := #_w1;
   IF #_w2 THEN "Tag_32" := TRUE; END_IF;
END_REGION

REGION Network 51
   RUNG wire#powerrail
      Contact( "FB11_DATA_ALARM_FB_DB".IW112.QH_ALM )
      wire#w1
      P_Trig( "DB9_P".P50 )
      S_Coil( "Tag_32" )
   END_RUNG
   RUNG wire#powerrail
      Contact( "FB11_DATA_ALARM_FB_DB".IW112.QL_ALM )
   END_RUNG wire#w1
   // the same network as SCL:
   #_w1 := "FB11_DATA_ALARM_FB_DB".IW112.QH_ALM OR "FB11_DATA_ALARM_FB_DB".IW112.QL_ALM;
   #_w2 := #_w1 AND NOT "DB9_P".P50;   // rising edge
   "DB9_P".P50 := #_w1;
   IF #_w2 THEN "Tag_32" := TRUE; END_IF;
END_REGION

REGION Network 52
   RUNG wire#powerrail
      Contact( "FB11_DATA_ALARM_FB_DB".IW114.QH_ALM )
      wire#w1
      P_Trig( "DB9_P".P51 )
      S_Coil( "Tag_32" )
   END_RUNG
   RUNG wire#powerrail
      Contact( "FB11_DATA_ALARM_FB_DB".IW114.QL_ALM )
   END_RUNG wire#w1
   // the same network as SCL:
   #_w1 := "FB11_DATA_ALARM_FB_DB".IW114.QH_ALM OR "FB11_DATA_ALARM_FB_DB".IW114.QL_ALM;
   #_w2 := #_w1 AND NOT "DB9_P".P51;   // rising edge
   "DB9_P".P51 := #_w1;
   IF #_w2 THEN "Tag_32" := TRUE; END_IF;
END_REGION

REGION Network 53
   RUNG wire#powerrail
      Contact( "FB11_DATA_ALARM_FB_DB".IW116.QH_ALM )
      wire#w1
      P_Trig( "DB9_P".P52 )
      S_Coil( "Tag_32" )
   END_RUNG
   RUNG wire#powerrail
      Contact( "FB11_DATA_ALARM_FB_DB".IW116.QL_ALM )
   END_RUNG wire#w1
   // the same network as SCL:
   #_w1 := "FB11_DATA_ALARM_FB_DB".IW116.QH_ALM OR "FB11_DATA_ALARM_FB_DB".IW116.QL_ALM;
   #_w2 := #_w1 AND NOT "DB9_P".P52;   // rising edge
   "DB9_P".P52 := #_w1;
   IF #_w2 THEN "Tag_32" := TRUE; END_IF;
END_REGION

REGION Network 54
   RUNG wire#powerrail
      Contact( "FB11_DATA_ALARM_FB_DB".PID400.QH_ALM )
      wire#w1
      P_Trig( "DB9_P".P53 )
      S_Coil( "Tag_32" )
   END_RUNG
   RUNG wire#powerrail
      Contact( "FB11_DATA_ALARM_FB_DB".PID400.QL_ALM )
   END_RUNG wire#w1
   // the same network as SCL:
   #_w1 := "FB11_DATA_ALARM_FB_DB".PID400.QH_ALM OR "FB11_DATA_ALARM_FB_DB".PID400.QL_ALM;
   #_w2 := #_w1 AND NOT "DB9_P".P53;   // rising edge
   "DB9_P".P53 := #_w1;
   IF #_w2 THEN "Tag_32" := TRUE; END_IF;
END_REGION

REGION Network 55
   RUNG wire#powerrail
      Contact( "FB11_DATA_ALARM_FB_DB".PID408.QH_ALM )
      wire#w1
      P_Trig( "DB9_P".P54 )
      S_Coil( "Tag_32" )
   END_RUNG
   RUNG wire#powerrail
      Contact( "FB11_DATA_ALARM_FB_DB".PID408.QL_ALM )
   END_RUNG wire#w1
   // the same network as SCL:
   #_w1 := "FB11_DATA_ALARM_FB_DB".PID408.QH_ALM OR "FB11_DATA_ALARM_FB_DB".PID408.QL_ALM;
   #_w2 := #_w1 AND NOT "DB9_P".P54;   // rising edge
   "DB9_P".P54 := #_w1;
   IF #_w2 THEN "Tag_32" := TRUE; END_IF;
END_REGION

REGION Network 56
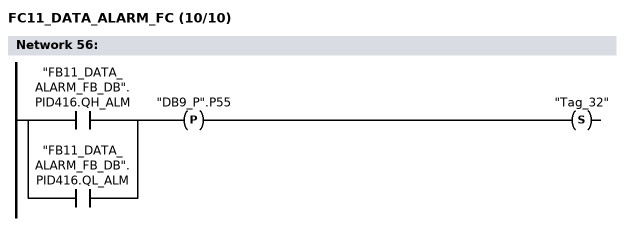
   RUNG wire#powerrail
      Contact( "FB11_DATA_ALARM_FB_DB".PID416.QH_ALM )
      wire#w1
      P_Trig( "DB9_P".P55 )
      S_Coil( "Tag_32" )
   END_RUNG
   RUNG wire#powerrail
      Contact( "FB11_DATA_ALARM_FB_DB".PID416.QL_ALM )
   END_RUNG wire#w1
   // the same network as SCL:
   #_w1 := "FB11_DATA_ALARM_FB_DB".PID416.QH_ALM OR "FB11_DATA_ALARM_FB_DB".PID416.QL_ALM;
   #_w2 := #_w1 AND NOT "DB9_P".P55;   // rising edge
   "DB9_P".P55 := #_w1;
   IF #_w2 THEN "Tag_32" := TRUE; END_IF;
END_REGION
END_FUNCTION

ORGANIZATION_BLOCK "Main"   // OB1, LAD, ProgramCycle
TITLE = "Main Program Sweep (Cycle)"
{ S7_Optimized_Access := 'TRUE' }
VERSION : 0.1
   VAR_INPUT
      Initial_Call : Bool;   // Initial call of this OB
      Remanence : Bool;   // =True, if remanent data are available
   END_VAR
BEGIN

REGION Network 1
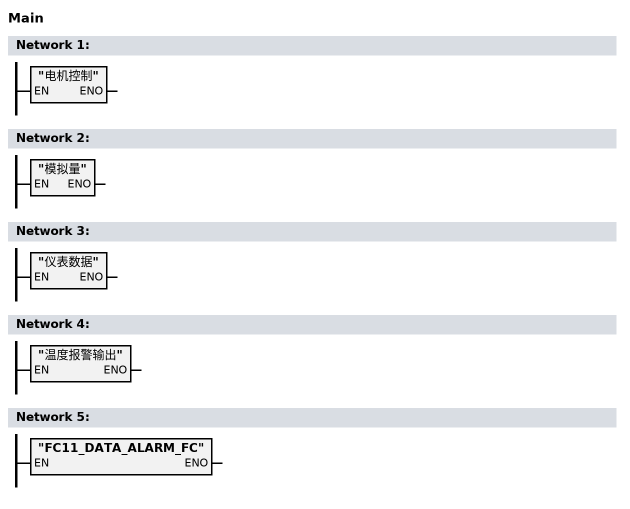
   RUNG wire#powerrail
      "电机控制"()
   END_RUNG
   // the same network as SCL:
   "电机控制"();
END_REGION

REGION Network 2
   RUNG wire#powerrail
      "模拟量"()
   END_RUNG
   // the same network as SCL:
   "模拟量"();
END_REGION

REGION Network 3
   RUNG wire#powerrail
      "仪表数据"()
   END_RUNG
   // the same network as SCL:
   "仪表数据"();
END_REGION

REGION Network 4
   RUNG wire#powerrail
      "温度报警输出"()
   END_RUNG
   // the same network as SCL:
   "温度报警输出"();
END_REGION

REGION Network 5
   RUNG wire#powerrail
      "FC11_DATA_ALARM_FC"()
   END_RUNG
   // the same network as SCL:
   "FC11_DATA_ALARM_FC"();
END_REGION
END_ORGANIZATION_BLOCK

ORGANIZATION_BLOCK "Cyclic interrupt"   // OB30, LAD, CyclicInterrupt
{ S7_Optimized_Access := 'TRUE' }
VERSION : 0.1
   VAR_INPUT
      Initial_Call : Bool;   // Initial call of this OB
      Event_Count : Int;   // Events discarded
   END_VAR
BEGIN

REGION Network 1
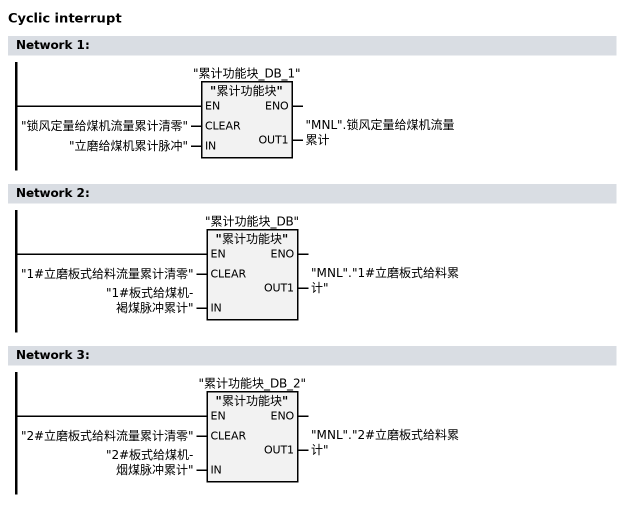
   RUNG wire#powerrail
      "累计功能块_DB_1"(CLEAR := "锁风定量给煤机流量累计清零", IN := "立磨给煤机累计脉冲", OUT1 => "MNL".锁风定量给煤机流量累计)
   END_RUNG
   // the same network as SCL:
   "累计功能块_DB_1"(CLEAR := "锁风定量给煤机流量累计清零", IN := "立磨给煤机累计脉冲", OUT1 => "MNL".锁风定量给煤机流量累计);   // "累计功能块"
END_REGION

REGION Network 2
   RUNG wire#powerrail
      "累计功能块_DB"(CLEAR := "1#立磨板式给料流量累计清零", IN := "1#板式给煤机-褐煤脉冲累计", OUT1 => "MNL"."1#立磨板式给料累计")
   END_RUNG
   // the same network as SCL:
   "累计功能块_DB"(CLEAR := "1#立磨板式给料流量累计清零", IN := "1#板式给煤机-褐煤脉冲累计", OUT1 => "MNL"."1#立磨板式给料累计");   // "累计功能块"
END_REGION

REGION Network 3
   RUNG wire#powerrail
      "累计功能块_DB_2"(CLEAR := "2#立磨板式给料流量累计清零", IN := "2#板式给煤机-烟煤脉冲累计", OUT1 => "MNL"."2#立磨板式给料累计")
   END_RUNG
   // the same network as SCL:
   "累计功能块_DB_2"(CLEAR := "2#立磨板式给料流量累计清零", IN := "2#板式给煤机-烟煤脉冲累计", OUT1 => "MNL"."2#立磨板式给料累计");   // "累计功能块"
END_REGION
END_ORGANIZATION_BLOCK